VERSION : 0.1
   VAR_INPUT
      Value : Real;
      "Raw Value" : Int;
      Enable : Bool := true;
      "Enable Delay Time" : Time := T#10s;
      "High Value Release" : Bool := true;   // It is Releasing High Values from Enable restriction
      "SHORT CIRCUIT VALUE" : Real := 32000.0;
      "BROKEN WIRE VALUE" : Real := -32000.0;
      "VERY LOW LEVEL VALUE (LL)" : Real;
      "LOW LEVEL VALUE (L)" : Real;
      "HIGH LEVEL VALUE (H)" : Real;
      "VERY HIGH LEVEL VALUE (HH)" : Real;
      OFFSET : Real;
      "ALARM DELAY" : Time := T#1s;
      "Peak Value Reset" : Bool;
   END_VAR
   VAR_OUTPUT
      "ALARM HH" : Bool;
      "ALARM H" : Bool;
      "ALARM L" : Bool;
      "ALARM LL" : Bool;
      "ALARM READING" : Bool;
      "Peak Value" : Real;
      Alarm : Word;
      Alarm_INT : Int;
   END_VAR
   VAR
      TRUE : Bool;
      FALSE : Bool;
      Raw_value_int : Int;
      RET_VAL : Word;
      RAW_scaled_mA : Real;
      RAW_scaled_VALUE : Real;
      SCALED_OFFSETTED_VALUE : Real;
      Error_present : Bool;
      "Enable Internal" : Bool;
      "ALARM HH_interm" : Bool;
      "ALARM H_interm" : Bool;
      "ALARM L_interm" : Bool;
      "ALARM LL_interm" : Bool;
      "ALARM READING_interm" : Bool;
      "ALARM_HH delay" : TON_TIME;
      "ALARM_H delay" : TON_TIME;
      "ALARM_LL delay" : TON_TIME;
      "ALARM_L delay" : TON_TIME;
      "ALARM_READING delay" : TON_TIME;
      "ALARM READING TOF" : TOF_TIME;
      "HI HI TOF" : TOF_TIME;
      "HI TOF" : TOF_TIME;
      "LOE TOF" : TOF_TIME;
      "LOW TOF" : TOF_TIME;
      "LOW LOW TOF" : TOF_TIME;
      "Enable TON" : TON_TIME;
   END_VAR
   VAR_TEMP   // added for the SCL form of the ladder/FBD networks
      _w1 : Bool;
   END_VAR
BEGIN

REGION Network 1: True False
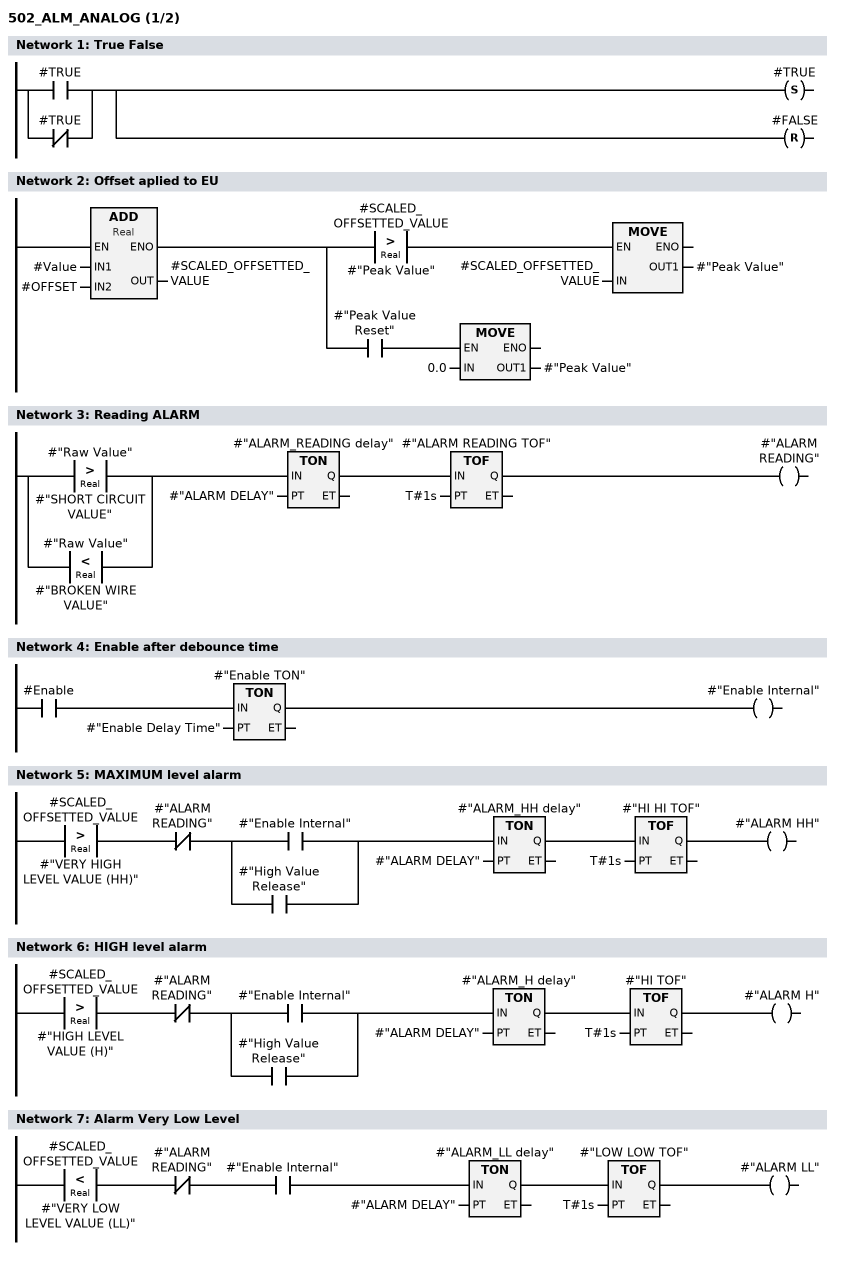
   RUNG wire#powerrail
      Contact( #TRUE )
      wire#w1
      S_Coil( #TRUE )
   END_RUNG
   RUNG wire#powerrail
      I_Contact( #TRUE )
   END_RUNG wire#w1
   RUNG wire#w1
      R_Coil( #FALSE )
   END_RUNG
   // the same network as SCL:
   #_w1 := #TRUE OR NOT #TRUE;
   IF #_w1 THEN
       #TRUE := TRUE;
       #FALSE := FALSE;
   END_IF;
END_REGION

REGION Network 2: Offset aplied to EU
   RUNG wire#powerrail
      { S7_Templates := "SrcType := Real"; S7_GenerateENO := "TRUE" } Add(in1 := #Value, in2 := #OFFSET, out => #SCALED_OFFSETTED_VALUE)
      wire#w1
      { S7_Templates := "SrcType := Real" } GT_Contact(in1 := #SCALED_OFFSETTED_VALUE, in2 := #"Peak Value")
      Move(in := #SCALED_OFFSETTED_VALUE, out1 => #"Peak Value")
   END_RUNG
   RUNG wire#w1
      Contact( #"Peak Value Reset" )
      Move(in := 0.0, out1 => #"Peak Value")
   END_RUNG
   // the same network as SCL:
   // ENO of a box is taken as its EN; it also drops when the box reports an error
   #SCALED_OFFSETTED_VALUE := #Value + #OFFSET;
   IF #SCALED_OFFSETTED_VALUE > #"Peak Value" THEN #"Peak Value" := #SCALED_OFFSETTED_VALUE; END_IF;
   IF #"Peak Value Reset" THEN #"Peak Value" := 0.0; END_IF;
END_REGION

REGION Network 3: Reading ALARM
   #"ALARM_READING delay"(IN := (#"Raw Value" > #"SHORT CIRCUIT VALUE") OR (#"Raw Value" < #"BROKEN WIRE VALUE"),   // TON
                          PT := #"ALARM DELAY");
   #"ALARM READING TOF"(IN := #"ALARM_READING delay".Q, PT := T#1s);   // TOF
   #"ALARM READING" := #"ALARM READING TOF".Q;
END_REGION

REGION Network 4: Enable after debounce time
   #"Enable TON"(IN := #Enable, PT := #"Enable Delay Time");   // TON
   #"Enable Internal" := #"Enable TON".Q;
END_REGION

REGION Network 5: MAXIMUM level alarm
   #"ALARM_HH delay"(IN := (#SCALED_OFFSETTED_VALUE > #"VERY HIGH LEVEL VALUE (HH)") AND NOT #"ALARM READING" AND (#"Enable Internal" OR #"High Value Release"),   // TON
                     PT := #"ALARM DELAY");
   #"HI HI TOF"(IN := #"ALARM_HH delay".Q, PT := T#1s);   // TOF
   #"ALARM HH" := #"HI HI TOF".Q;
END_REGION

REGION Network 6: HIGH level alarm
   #"ALARM_H delay"(IN := (#SCALED_OFFSETTED_VALUE > #"HIGH LEVEL VALUE (H)") AND NOT #"ALARM READING" AND (#"Enable Internal" OR #"High Value Release"),   // TON
                    PT := #"ALARM DELAY");
   #"HI TOF"(IN := #"ALARM_H delay".Q, PT := T#1s);   // TOF
   #"ALARM H" := #"HI TOF".Q;
END_REGION

REGION Network 7: Alarm Very Low Level
   #"ALARM_LL delay"(IN := (#SCALED_OFFSETTED_VALUE < #"VERY LOW LEVEL VALUE (LL)") AND NOT #"ALARM READING" AND #"Enable Internal",   // TON
                     PT := #"ALARM DELAY");
   #"LOW LOW TOF"(IN := #"ALARM_LL delay".Q, PT := T#1s);   // TOF
   #"ALARM LL" := #"LOW LOW TOF".Q;
END_REGION

REGION Network 8: Alarm Low Level
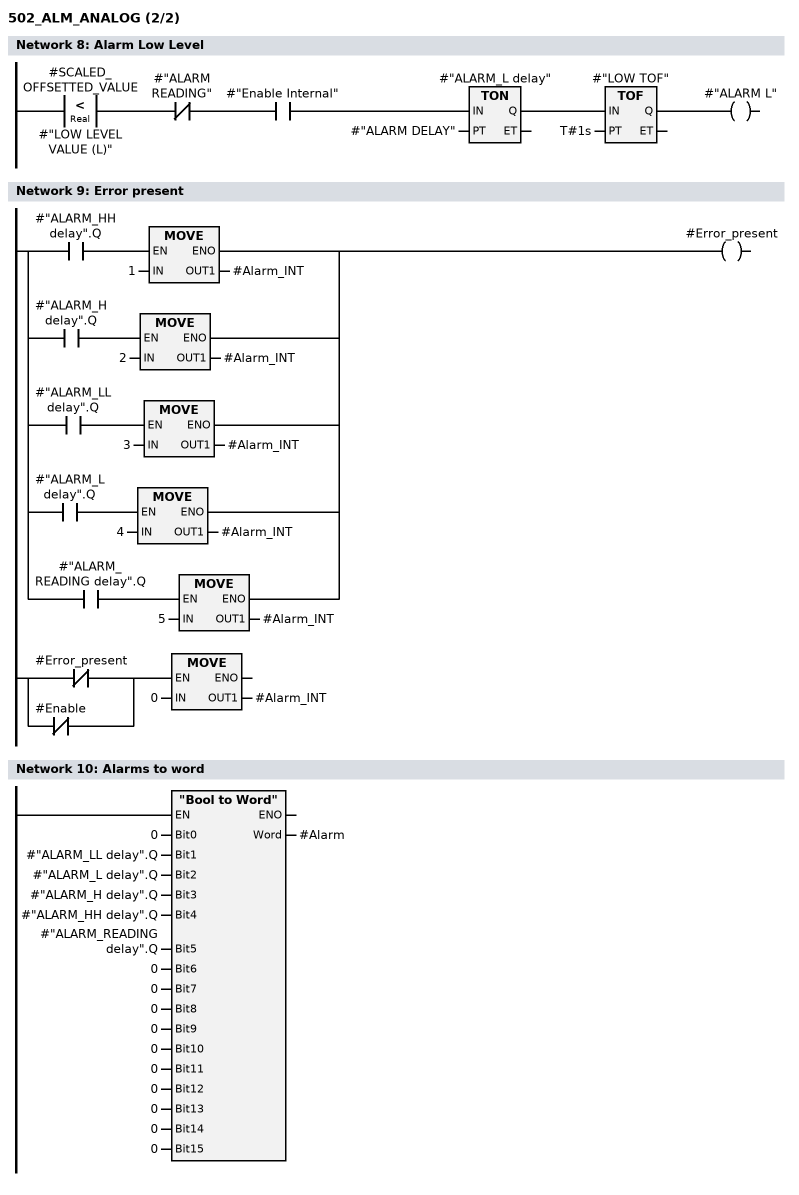
   #"ALARM_L delay"(IN := (#SCALED_OFFSETTED_VALUE < #"LOW LEVEL VALUE (L)") AND NOT #"ALARM READING" AND #"Enable Internal",   // TON
                    PT := #"ALARM DELAY");
   #"LOW TOF"(IN := #"ALARM_L delay".Q, PT := T#1s);   // TOF
   #"ALARM L" := #"LOW TOF".Q;
END_REGION

REGION Network 9: Error present
   RUNG wire#powerrail
      Contact( #"ALARM_HH delay".Q )
      { S7_GenerateENO := "TRUE" } Move(in := 1, out1 => #Alarm_INT)
      wire#w1
      Coil( #Error_present )
   END_RUNG
   RUNG wire#powerrail
      Contact( #"ALARM_H delay".Q )
      { S7_GenerateENO := "TRUE" } Move(in := 2, out1 => #Alarm_INT)
   END_RUNG wire#w1
   RUNG wire#powerrail
      Contact( #"ALARM_LL delay".Q )
      { S7_GenerateENO := "TRUE" } Move(in := 3, out1 => #Alarm_INT)
   END_RUNG wire#w1
   RUNG wire#powerrail
      Contact( #"ALARM_L delay".Q )
      { S7_GenerateENO := "TRUE" } Move(in := 4, out1 => #Alarm_INT)
   END_RUNG wire#w1
   RUNG wire#powerrail
      Contact( #"ALARM_READING delay".Q )
      { S7_GenerateENO := "TRUE" } Move(in := 5, out1 => #Alarm_INT)
   END_RUNG wire#w1
   RUNG wire#powerrail
      I_Contact( #Error_present )
      wire#w2
      Move(in := 0, out1 => #Alarm_INT)
   END_RUNG
   RUNG wire#powerrail
      I_Contact( #Enable )
   END_RUNG wire#w2
   // the same network as SCL:
   // ENO of a box is taken as its EN; it also drops when the box reports an error
   IF #"ALARM_HH delay".Q THEN #Alarm_INT := 1; END_IF;
   IF #"ALARM_H delay".Q THEN #Alarm_INT := 2; END_IF;
   IF #"ALARM_LL delay".Q THEN #Alarm_INT := 3; END_IF;
   IF #"ALARM_L delay".Q THEN #Alarm_INT := 4; END_IF;
   IF #"ALARM_READING delay".Q THEN #Alarm_INT := 5; END_IF;
   #Error_present := #"ALARM_HH delay".Q OR #"ALARM_H delay".Q OR #"ALARM_LL delay".Q OR #"ALARM_L delay".Q OR #"ALARM_READING delay".Q;
   IF NOT #Error_present OR NOT #Enable THEN #Alarm_INT := 0; END_IF;
END_REGION

REGION Network 10: Alarms to word
   RUNG wire#powerrail
      "Bool to Word"(Bit0 := 0, Bit1 := #"ALARM_LL delay".Q, Bit2 := #"ALARM_L delay".Q, Bit3 := #"ALARM_H delay".Q, Bit4 := #"ALARM_HH delay".Q, Bit5 := #"ALARM_READING delay".Q, Bit6 := 0, Bit7 := 0, Bit8 := 0, Bit9 := 0, Bit10 := 0, Bit11 := 0, Bit12 := 0, Bit13 := 0, Bit14 := 0, Bit15 := 0, "Word" => #Alarm)
   END_RUNG
   // the same network as SCL:
   "Bool to Word"(Bit0 := 0,
                  Bit1 := #"ALARM_LL delay".Q,
                  Bit2 := #"ALARM_L delay".Q,
                  Bit3 := #"ALARM_H delay".Q,
                  Bit4 := #"ALARM_HH delay".Q,
                  Bit5 := #"ALARM_READING delay".Q,
                  Bit6 := 0,
                  Bit7 := 0,
                  Bit8 := 0,
                  Bit9 := 0,
                  Bit10 := 0,
                  Bit11 := 0,
                  Bit12 := 0,
                  Bit13 := 0,
                  Bit14 := 0,
                  Bit15 := 0,
                  "Word" => #Alarm);
END_REGION
END_FUNCTION_BLOCK

FUNCTION_BLOCK "503_ALARM CHCK"   // FB503, LAD
{ S7_Optimized_Access := 'TRUE' }
VERSION : 0.1
   VAR_INPUT
      "Alarm Word 1" : Word;
      "Alarm Word 2" : Word;
      "Alarm Word 3" : Word;
      "Alarm Word 4" : Word;
      "Alarm Word 5" : Word;
      "Alarm Word 6" : Word;
      "Alarm Word 7" : Word;
      "Alarm Word 8" : Word;
      "Alarm Word 9" : Word;
      "Alarm Word 10" : Word;
      "Alarm Word 11" : Word;
      "Alarm Word 12" : Word;
      "Alarm Word 13" : Word;
      "Alarm Word 14" : Word;
      "Alarm Word 15" : Word;
      "Alarm Word 16" : Word;
      "Reset Alarm" : Bool;
   END_VAR
   VAR_OUTPUT
      "Sound Alarm" : Bool;
   END_VAR
   VAR
      "Alarm Word Interm 1" : Word;
      "Alarm Word Interm 2" : Word;
      "Alarm Word Interm 3" : Word;
      "Alarm Word Interm 4" : Word;
      "Alarm Word Interm 5" : Word;
      "Alarm Word Interm 6" : Word;
      "Alarm Word Interm 7" : Word;
      "Alarm Word Interm 8" : Word;
      "Alarm Word Interm 9" : Word;
      "Alarm Word Interm 10" : Word;
      "Alarm Word Interm 11" : Word;
      "Alarm Word Interm 12" : Word;
      "Alarm Word Interm 13" : Word;
      "Alarm Word Interm 14" : Word;
      "Alarm Word Interm 15" : Word;
      "Alarm Word Interm 16" : Word;
      "Alarm Word bool 1" : Bool;
      "Alarm Word bool 2" : Bool;
      "Alarm Word bool 3" : Bool;
      "Alarm Word bool 4" : Bool;
      "Alarm Word bool 5" : Bool;
      "Alarm Word bool 6" : Bool;
      "Alarm Word bool 7" : Bool;
      "Alarm Word bool 8" : Bool;
      "Alarm Word bool 9" : Bool;
      "Alarm Word bool 10" : Bool;
      "Alarm Word bool 11" : Bool;
      "Alarm Word bool 12" : Bool;
      "Alarm Word bool 13" : Bool;
      "Alarm Word bool 14" : Bool;
      "Alarm Word bool 15" : Bool;
      "Alarm Word bool 16" : Bool;
      "Delayed Alarm Reset" : TON_TIME;
   END_VAR
BEGIN

REGION Network 1: Check Words
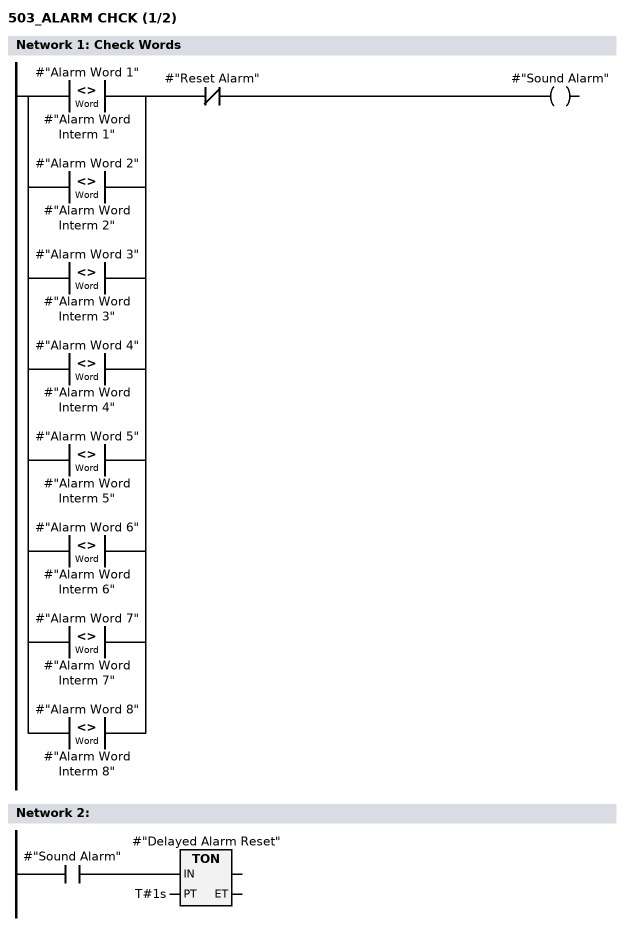
   RUNG wire#powerrail
      { S7_Templates := "SrcType := Word" } NE_Contact(in1 := #"Alarm Word 1", in2 := #"Alarm Word Interm 1")
      wire#w1
      I_Contact( #"Reset Alarm" )
      Coil( #"Sound Alarm" )
   END_RUNG
   RUNG wire#powerrail
      { S7_Templates := "SrcType := Word" } NE_Contact(in1 := #"Alarm Word 2", in2 := #"Alarm Word Interm 2")
   END_RUNG wire#w1
   RUNG wire#powerrail
      { S7_Templates := "SrcType := Word" } NE_Contact(in1 := #"Alarm Word 3", in2 := #"Alarm Word Interm 3")
   END_RUNG wire#w1
   RUNG wire#powerrail
      { S7_Templates := "SrcType := Word" } NE_Contact(in1 := #"Alarm Word 4", in2 := #"Alarm Word Interm 4")
   END_RUNG wire#w1
   RUNG wire#powerrail
      { S7_Templates := "SrcType := Word" } NE_Contact(in1 := #"Alarm Word 5", in2 := #"Alarm Word Interm 5")
   END_RUNG wire#w1
   RUNG wire#powerrail
      { S7_Templates := "SrcType := Word" } NE_Contact(in1 := #"Alarm Word 6", in2 := #"Alarm Word Interm 6")
   END_RUNG wire#w1
   RUNG wire#powerrail
      { S7_Templates := "SrcType := Word" } NE_Contact(in1 := #"Alarm Word 7", in2 := #"Alarm Word Interm 7")
   END_RUNG wire#w1
   RUNG wire#powerrail
      { S7_Templates := "SrcType := Word" } NE_Contact(in1 := #"Alarm Word 8", in2 := #"Alarm Word Interm 8")
   END_RUNG wire#w1
   // the same network as SCL:
   #"Sound Alarm" := ((#"Alarm Word 1" <> #"Alarm Word Interm 1") OR (#"Alarm Word 2" <> #"Alarm Word Interm 2") OR (#"Alarm Word 3" <> #"Alarm Word Interm 3") OR (#"Alarm Word 4" <> #"Alarm Word Interm 4") OR (#"Alarm Word 5" <> #"Alarm Word Interm 5") OR (#"Alarm Word 6" <> #"Alarm Word Interm 6") OR (#"Alarm Word 7" <> #"Alarm Word Interm 7") OR (#"Alarm Word 8" <> #"Alarm Word Interm 8")) AND NOT #"Reset Alarm";
END_REGION

REGION Network 2
   #"Delayed Alarm Reset"(IN := #"Sound Alarm", PT := T#1s);   // TON
END_REGION

REGION Network 3: Move Words
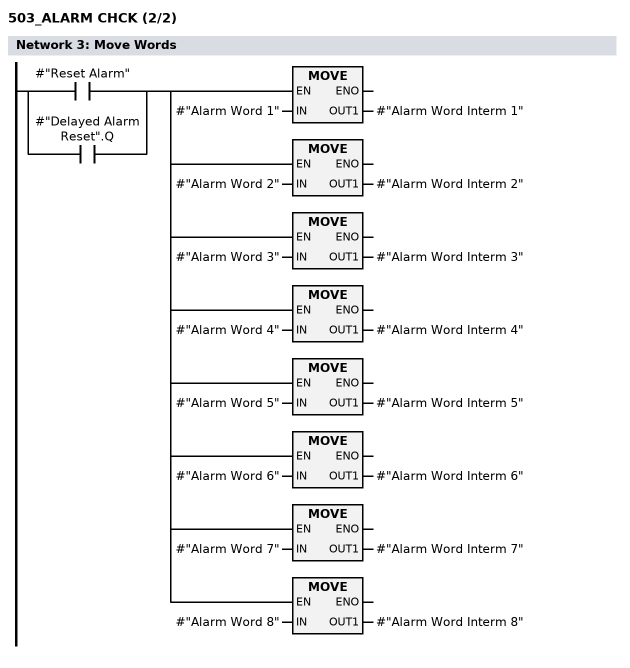
   RUNG wire#powerrail
      Contact( #"Reset Alarm" )
      wire#w1
      Move(in := #"Alarm Word 1", out1 => #"Alarm Word Interm 1")
   END_RUNG
   RUNG wire#powerrail
      Contact( #"Delayed Alarm Reset".Q )
   END_RUNG wire#w1
   RUNG wire#w1
      Move(in := #"Alarm Word 2", out1 => #"Alarm Word Interm 2")
   END_RUNG
   RUNG wire#w1
      Move(in := #"Alarm Word 3", out1 => #"Alarm Word Interm 3")
   END_RUNG
   RUNG wire#w1
      Move(in := #"Alarm Word 4", out1 => #"Alarm Word Interm 4")
   END_RUNG
   RUNG wire#w1
      Move(in := #"Alarm Word 5", out1 => #"Alarm Word Interm 5")
   END_RUNG
   RUNG wire#w1
      Move(in := #"Alarm Word 6", out1 => #"Alarm Word Interm 6")
   END_RUNG
   RUNG wire#w1
      Move(in := #"Alarm Word 7", out1 => #"Alarm Word Interm 7")
   END_RUNG
   RUNG wire#w1
      Move(in := #"Alarm Word 8", out1 => #"Alarm Word Interm 8")
   END_RUNG
   // the same network as SCL:
   IF #"Reset Alarm" OR #"Delayed Alarm Reset".Q THEN
       #"Alarm Word Interm 1" := #"Alarm Word 1";
       #"Alarm Word Interm 2" := #"Alarm Word 2";
       #"Alarm Word Interm 3" := #"Alarm Word 3";
       #"Alarm Word Interm 4" := #"Alarm Word 4";
       #"Alarm Word Interm 5" := #"Alarm Word 5";
       #"Alarm Word Interm 6" := #"Alarm Word 6";
       #"Alarm Word Interm 7" := #"Alarm Word 7";
       #"Alarm Word Interm 8" := #"Alarm Word 8";
   END_IF;
END_REGION
END_FUNCTION_BLOCK

FUNCTION_BLOCK "Animation"   // FB515, LAD
{ S7_Optimized_Access := 'TRUE' }
VERSION : 0.1
   VAR_INPUT
      Run : Bool;
      Revert : Bool := true;
      "States Number" : Int := 10;
      Period : Time := T#250ms;
   END_VAR
   VAR_OUTPUT
      Animation : Int;
   END_VAR
   VAR RETAIN
      "Animation State" : CTU_INT;
      Reset : Bool;
   END_VAR
   VAR
      "Revert Aux" : Bool;
      LD : Bool;
      OFF : TON_TIME;
      ON : TON_TIME;
   END_VAR
BEGIN

REGION Network 1
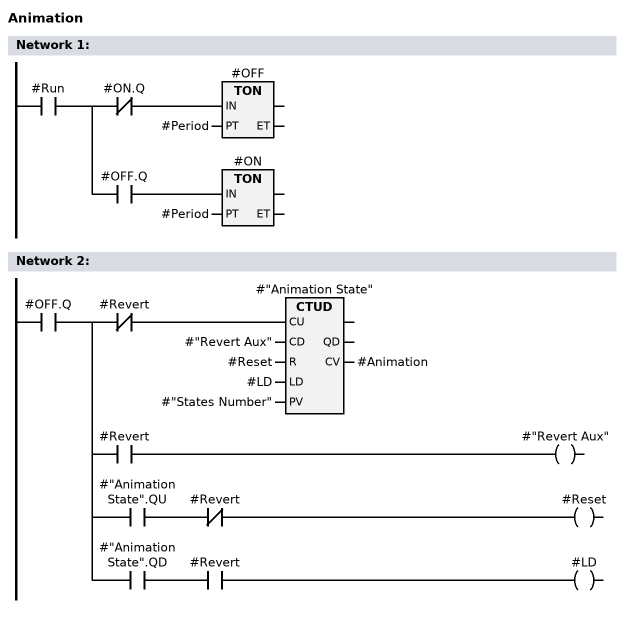
   #OFF(IN := #Run AND NOT #ON.Q, PT := #Period);   // TON
   #ON(IN := #Run AND #OFF.Q, PT := #Period);   // TON
END_REGION

REGION Network 2
   #"Animation State"(CU := #OFF.Q AND NOT #Revert,   // CTUD
                      CD := #"Revert Aux",
                      R := #Reset,
                      LD := #LD,
                      PV := #"States Number",
                      CV => #Animation);
   #"Revert Aux" := #OFF.Q AND #Revert;
   #Reset := #OFF.Q AND #"Animation State".QU AND NOT #Revert;
   #LD := #OFF.Q AND #"Animation State".QD AND #Revert;
END_REGION
END_FUNCTION_BLOCK

FUNCTION "Bool to Word" : Void   // FC202, FBD
{ S7_Optimized_Access := 'FALSE' }
VERSION : 0.1
// Die Funktion gruppiert 16 Variablen vom Datentyp "Bool" zu einer Variablen vom Datentyp "Word".
// *******************************************************************************
// The function groups 16 variables with type of data "Bool" to a variable with type of data "Word".
   VAR_INPUT
      Bit0 : Bool;
      Bit1 : Bool;
      Bit2 : Bool;
      Bit3 : Bool;
      Bit4 : Bool;
      Bit5 : Bool;
      Bit6 : Bool;
      Bit7 : Bool;
      Bit8 : Bool;
      Bit9 : Bool;
      Bit10 : Bool;
      Bit11 : Bool;
      Bit12 : Bool;
      Bit13 : Bool;
      Bit14 : Bool;
      Bit15 : Bool;
   END_VAR
   VAR_OUTPUT
      "Word" : Word;
   END_VAR
   VAR_TEMP
      aux : DInt;
   END_VAR
BEGIN

REGION Network 1: aux
   // Setze Hilfsvariable "aux" auf den Anfangswert 0.
   // ***************************************************************************
   // Set the auxiliary variable "aux" to the initial value 0.
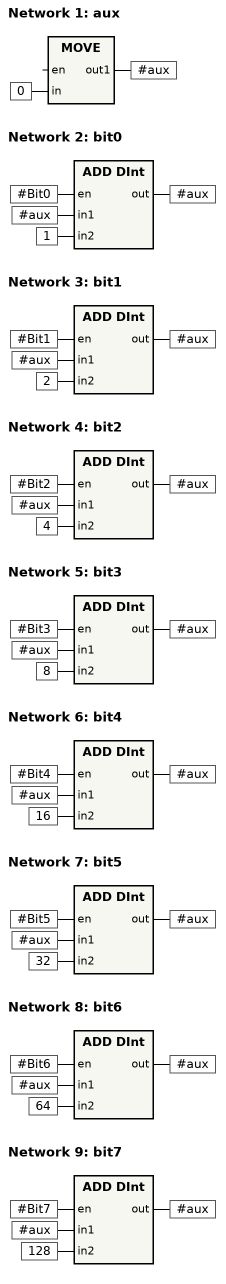
   #aux := 0;
END_REGION

REGION Network 2: bit0
   // Addiere Bit 0 zur Hilfsvariable "aux" vom Datentyp "UInt".
   // ***************************************************************************
   // Add Bit 0 to the auxiliary variable "aux" with type of data "UInt".
   IF #Bit0 THEN #aux := #aux + 1; END_IF;
END_REGION

REGION Network 3: bit1
   // Addiere Bit 1 zur Hilfsvariable "aux".
   // ***************************************************************************
   // Add Bit 1 to the auxiliary variable "aux".
   IF #Bit1 THEN #aux := #aux + 2; END_IF;
END_REGION

REGION Network 4: bit2
   // Addiere Bit 2 zur Hilfsvariable "aux".
   // ***************************************************************************
   // Add Bit 2 to the auxiliary variable "aux".
   IF #Bit2 THEN #aux := #aux + 4; END_IF;
END_REGION

REGION Network 5: bit3
   // Addiere Bit 3 zur Hilfsvariable "aux".
   // ***************************************************************************
   // Add Bit 3 to the auxiliary variable "aux".
   IF #Bit3 THEN #aux := #aux + 8; END_IF;
END_REGION

REGION Network 6: bit4
   // Addiere Bit 4 zur Hilfsvariable "aux".
   // ***************************************************************************
   // Add Bit 4 to the auxiliary variable "aux".
   IF #Bit4 THEN #aux := #aux + 16; END_IF;
END_REGION

REGION Network 7: bit5
   // Addiere Bit 5 zur Hilfsvariable "aux".
   // ***************************************************************************
   // Add Bit 5 to the auxiliary variable "aux".
   IF #Bit5 THEN #aux := #aux + 32; END_IF;
END_REGION

REGION Network 8: bit6
   // Addiere Bit 6 zur Hilfsvariable "aux".
   // ***************************************************************************
   // Add Bit 6 to the auxiliary variable "aux".
   IF #Bit6 THEN #aux := #aux + 64; END_IF;
END_REGION

REGION Network 9: bit7
   // Addiere Bit 7 zur Hilfsvariable "aux".
   // ***************************************************************************
   // Add Bit 7 to the auxiliary variable "aux".
   IF #Bit7 THEN #aux := #aux + 128; END_IF;
END_REGION

REGION Network 10: bit8
   // Addiere Bit 8 zur Hilfsvariable "aux".
   // ***************************************************************************
   // Add Bit 8 to the auxiliary variable "aux".
